        rgtTrkConv[6].Cap[0].dCenterPosConv_cmm := 258800, rgtTrkConv[6].Cap[0].dHeadPos_cmm := 2015800, rgtTrkConv[6].Cap[0].dHeadPosConv_cmm := 388800, rgtTrkConv[6].Cap[0].dPresenceHead_cmm := 2015800, rgtTrkConv[6].Cap[0].dPresenceTail_cmm := 1755800, rgtTrkConv[7].xGlassPresence := 1, rgtTrkConv[7].xPlatePassageNext := 1, rgtTrkConv[7].xGlassPresCom := 1, rgtTrkConv[7].xHeadPresenceConv := 1, rgtTrkConv[7].dStartPosition_cmm := 2127000, rgtTrkConv[7].dEndPosition_cmm := 2627000, rgtTrkConv[7].dStepAdv_cmm[0] := 1620, rgtTrkConv[7].dActualRamp_cmm[0] := 33700, rgtTrkConv[7].dLengthConveyor := 500000, rgtTrkConv[7].dHeadPosition_cmm := 2613400, rgtTrkConv[7].dTailPosition_cmm := 2445700, rgtTrkConv[7].dIndexCaps := 1, rgtTrkConv[7].Cap[0].xHead := 1, rgtTrkConv[7].Cap[0].xCenter := 1, rgtTrkConv[7].Cap[0].xTail := 1, rgtTrkConv[7].Cap[0].xPresence := 1, rgtTrkConv[7].Cap[0].dPointer := 12, rgtTrkConv[7].Cap[0].dTailPos_cmm := 2445700, rgtTrkConv[7].Cap[0].dTailPosConv_cmm := 318700, rgtTrkConv[7].Cap[0].dCenterPos_cmm := 2529550, rgtTrkConv[7].Cap[0].dCenterPosConv_cmm := 402550, rgtTrkConv[7].Cap[0].dHeadPos_cmm := 2613400, rgtTrkConv[7].Cap[0].dHeadPosConv_cmm := 486400, rgtTrkConv[7].Cap[0].dPresenceHead_cmm := 2613400, rgtTrkConv[7].Cap[0].dPresenceTail_cmm := 2445700, rgtTrkConv[8].xPlatePassagePrevious := 1, rgtTrkConv[8].xGlassPresCom := 1, rgtTrkConv[8].dStartPosition_cmm := 2627000, rgtTrkConv[8].dEndPosition_cmm := 2702000, rgtTrkConv[8].dStepAdv_cmm[0] := 1620, rgtTrkConv[8].dActualRamp_cmm[0] := 33700, rgtTrkConv[8].dLengthConveyor := 75000, rgtTrkConv[9].dStartPosition_cmm := 2702000, rgtTrkConv[9].dEndPosition_cmm := 3027000, rgtTrkConv[9].dStepAdv_cmm[0] := 2355, rgtTrkConv[9].dActualRamp_cmm[0] := 33700, rgtTrkConv[9].dLengthConveyor := 325000, rgtTrkConv[10].xGlassPresence := 1, rgtTrkConv[10].xGlassPresCom := 1, rgtTrkConv[10].xHeadPresenceConv := 1, rgtTrkConv[10].dStartPosition_cmm := 3027000, rgtTrkConv[10].dEndPosition_cmm := 3427000, rgtTrkConv[10].dStepAdv_cmm[0] := 2700, rgtTrkConv[10].dActualRamp_cmm[0] := 93700, rgtTrkConv[10].dLengthConveyor := 400000, rgtTrkConv[10].dHeadPosition_cmm := 3312224, rgtTrkConv[10].dTailPosition_cmm := 3052224, rgtTrkConv[10].dIndexCaps := 1, rgtTrkConv[10].Cap[0].xHead := 1, rgtTrkConv[10].Cap[0].xCenter := 1, rgtTrkConv[10].Cap[0].xTail := 1, rgtTrkConv[10].Cap[0].xPresence := 1, rgtTrkConv[10].Cap[0].dPointer := 1, rgtTrkConv[10].Cap[0].dTailPos_cmm := 3052224, rgtTrkConv[10].Cap[0].dTailPosConv_cmm := 25224,
        rgtTrkConv[10].Cap[0].dCenterPos_cmm := 3182224, rgtTrkConv[10].Cap[0].dCenterPosConv_cmm := 155224, rgtTrkConv[10].Cap[0].dHeadPos_cmm := 3312224, rgtTrkConv[10].Cap[0].dHeadPosConv_cmm := 285224, rgtTrkConv[10].Cap[0].dPresenceHead_cmm := 3312224, rgtTrkConv[10].Cap[0].dPresenceTail_cmm := 3052224, rgtTrkConv[11].dStartPosition_cmm := 3427000, rgtTrkConv[11].dEndPosition_cmm := 3777000, rgtTrkConv[11].dStepAdv_cmm[0] := 3000, rgtTrkConv[11].dStepAdv_cmm[1] := 3000, rgtTrkConv[11].dActualRamp_cmm[0] := 93700, rgtTrkConv[11].dActualRamp_cmm[1] := 93700, rgtTrkConv[11].dLengthConveyor := 350000, rgtTrkConv[12].xGlassPresence := 1, rgtTrkConv[12].xPlatePassageNext := 1, rgtTrkConv[12].xGlassPresCom := 1, rgtTrkConv[12].dStartPosition_cmm := 3777000, rgtTrkConv[12].dEndPosition_cmm := 4227000, rgtTrkConv[12].dStepAdv_cmm[0] := 3000, rgtTrkConv[12].dActualRamp_cmm[0] := 93700, rgtTrkConv[12].dLengthConveyor := 450000, rgtTrkConv[12].dTailPosition_cmm := 4202979, rgtTrkConv[12].dIndexCaps := 1, rgtTrkConv[12].Cap[0].xTail := 1, rgtTrkConv[12].Cap[0].xPresence := 1, rgtTrkConv[12].Cap[0].dPointer := 3, rgtTrkConv[12].Cap[0].dTailPos_cmm := 4202979, rgtTrkConv[12].Cap[0].dTailPosConv_cmm := 425979, rgtTrkConv[12].Cap[0].dPresenceHead_cmm := 4370679, rgtTrkConv[12].Cap[0].dPresenceTail_cmm := 4202979, rgtTrkConv[13].xGlassPresence := 1, rgtTrkConv[13].xPlatePassagePrevious := 1, rgtTrkConv[13].xGlassPresCom := 1, rgtTrkConv[13].xHeadPresenceConv := 1, rgtTrkConv[13].dStartPosition_cmm := 4227000, rgtTrkConv[13].dEndPosition_cmm := 4527000, rgtTrkConv[13].dStepAdv_cmm[0] := 3000, rgtTrkConv[13].dStepAdv_cmm[1] := 3000, rgtTrkConv[13].dActualRamp_cmm[0] := 93700, rgtTrkConv[13].dActualRamp_cmm[1] := 93700, rgtTrkConv[13].dLengthConveyor := 300000, rgtTrkConv[13].dHeadPosition_cmm := 4370679, rgtTrkConv[13].dIndexCaps := 1, rgtTrkConv[13].Cap[0].xHead := 1, rgtTrkConv[13].Cap[0].xCenter := 1, rgtTrkConv[13].Cap[0].xPresence := 1, rgtTrkConv[13].Cap[0].dPointer := 3, rgtTrkConv[13].Cap[0].dCenterPos_cmm := 4286829, rgtTrkConv[13].Cap[0].dCenterPosConv_cmm := 59829, rgtTrkConv[13].Cap[0].dHeadPos_cmm := 4370679, rgtTrkConv[13].Cap[0].dHeadPosConv_cmm := 143679, rgtTrkConv[13].Cap[0].dPresenceHead_cmm := 4370679, rgtTrkConv[13].Cap[0].dPresenceTail_cmm := 4202979, rgtTrkConv[14].dStartPosition_cmm := 4527000, rgtTrkConv[14].dEndPosition_cmm := 4627000, rgtTrkConv[14].dStepAdv_cmm[0] := 3300, rgtTrkConv[14].dStepAdv_cmm[1] := 3300, rgtTrkConv[14].dActualRamp_cmm[0] := 93700, rgtTrkConv[14].dActualRamp_cmm[1] := 93700, rgtTrkConv[14].dLengthConveyor := 100000,
        rgtTrkConv[15].dStartPosition_cmm := 4627000, rgtTrkConv[15].dEndPosition_cmm := 5027000, rgtTrkConv[15].dStepAdv_cmm[0] := 2514, rgtTrkConv[15].dActualRamp_cmm[0] := 93700, rgtTrkConv[15].dLengthConveyor := 400000, rgtTrkConv[15].tmON_StopNextConveyor.PRE := 20, rgtTrkConv[16].dStartPosition_cmm := 5027000, rgtTrkConv[16].dEndPosition_cmm := 5427000, rgtTrkConv[16].dStepAdv_cmm[0] := 3300, rgtTrkConv[16].dActualRamp_cmm[0] := 93700, rgtTrkConv[16].dLengthConveyor := 400000, rgtTrkConv[17].dStartPosition_cmm := 5427000, rgtTrkConv[17].dEndPosition_cmm := 5827000, rgtTrkConv[17].dStepAdv_cmm[0] := 2700, rgtTrkConv[17].dActualRamp_cmm[0] := 93700, rgtTrkConv[17].dLengthConveyor := 400000, rgtTrkConv[18].xGlassPresence := 1, rgtTrkConv[18].xPlatePassageNext := 1, rgtTrkConv[18].xGlassPresCom := 1, rgtTrkConv[18].dStartPosition_cmm := 5827000, rgtTrkConv[18].dEndPosition_cmm := 6227000, rgtTrkConv[18].dStepAdv_cmm[0] := 2700, rgtTrkConv[18].dStepAdv_cmm[1] := 2700, rgtTrkConv[18].dActualRamp_cmm[0] := 93700, rgtTrkConv[18].dActualRamp_cmm[1] := 93700, rgtTrkConv[18].dLengthConveyor := 400000, rgtTrkConv[18].dTailPosition_cmm := 6128300, rgtTrkConv[18].dIndexCaps := 1, rgtTrkConv[18].Cap[0].xCenter := 1, rgtTrkConv[18].Cap[0].xTail := 1, rgtTrkConv[18].Cap[0].xPresence := 1, rgtTrkConv[18].Cap[0].dPointer := 8, rgtTrkConv[18].Cap[0].dTailPos_cmm := 6128300, rgtTrkConv[18].Cap[0].dTailPosConv_cmm := 301300, rgtTrkConv[18].Cap[0].dCenterPos_cmm := 6212150, rgtTrkConv[18].Cap[0].dCenterPosConv_cmm := 385150, rgtTrkConv[18].Cap[0].dPresenceHead_cmm := 6296000, rgtTrkConv[18].Cap[0].dPresenceTail_cmm := 6128300, rgtTrkConv[19].xGlassPresence := 1, rgtTrkConv[19].xPlatePassagePrevious := 1, rgtTrkConv[19].xGlassPresCom := 1, rgtTrkConv[19].xHeadPresenceConv := 1, rgtTrkConv[19].dStartPosition_cmm := 6227000, rgtTrkConv[19].dEndPosition_cmm := 6627000, rgtTrkConv[19].dStepAdv_cmm[0] := 2700, rgtTrkConv[19].dActualRamp_cmm[0] := 93700, rgtTrkConv[19].dLengthConveyor := 400000, rgtTrkConv[19].dHeadPosition_cmm := 6296000, rgtTrkConv[19].dIndexCaps := 1, rgtTrkConv[19].Cap[0].xHead := 1, rgtTrkConv[19].Cap[0].xPresence := 1, rgtTrkConv[19].Cap[0].dPointer := 8, rgtTrkConv[19].Cap[0].dHeadPos_cmm := 6296000, rgtTrkConv[19].Cap[0].dHeadPosConv_cmm := 69000, rgtTrkConv[19].Cap[0].dPresenceHead_cmm := 6296000, rgtTrkConv[19].Cap[0].dPresenceTail_cmm := 6128300, rgtTrkConv[20].dStartPosition_cmm := 6627000, rgtTrkConv[20].dEndPosition_cmm := 7027000, rgtTrkConv[20].dStepAdv_cmm[0] := 2700, rgtTrkConv[20].dActualRamp_cmm[0] := 93700,
        rgtTrkConv[20].dLengthConveyor := 400000, rgtTrkConv[21].dStartPosition_cmm := 7027000, rgtTrkConv[21].dEndPosition_cmm := 7427000, rgtTrkConv[21].dStepAdv_cmm[0] := 87, rgtTrkConv[21].dActualRamp_cmm[0] := 93700, rgtTrkConv[21].dLengthConveyor := 400000, rgtTrkConv[22].dStartPosition_cmm := 7427000, rgtTrkConv[22].dEndPosition_cmm := 8177000, rgtTrkConv[22].dStepAdv_cmm[0] := 3000, rgtTrkConv[22].dActualRamp_cmm[0] := 93700, rgtTrkConv[22].dLengthConveyor := 750000, rgtTrkConv[23].dStartPosition_cmm := 8177000, rgtTrkConv[23].dEndPosition_cmm := 8627000, rgtTrkConv[23].dStepAdv_cmm[0] := 3000, rgtTrkConv[23].dActualRamp_cmm[0] := 93700, rgtTrkConv[23].dLengthConveyor := 450000, rgtTrkConv[24].dStartPosition_cmm := 8627000, rgtTrkConv[24].dEndPosition_cmm := 9077000, rgtTrkConv[24].dStepAdv_cmm[0] := 3300, rgtTrkConv[24].dActualRamp_cmm[0] := 93700, rgtTrkConv[24].dLengthConveyor := 450000, rgtTrkConv[25].dStartPosition_cmm := 9077000, rgtTrkConv[25].dEndPosition_cmm := 9372000, rgtTrkConv[25].dStepAdv_cmm[0] := 3300, rgtTrkConv[25].dActualRamp_cmm[0] := 93700, rgtTrkConv[25].dLengthConveyor := 295000, rgtTrkConv[25].tmON_StopNextConveyor.PRE := 20, rgtTrkConv[26].dStartPosition_cmm := 9372000, rgtTrkConv[26].dEndPosition_cmm := 9897000, rgtTrkConv[26].dStepAdv_cmm[0] := 3300, rgtTrkConv[26].dActualRamp_cmm[0] := 93700, rgtTrkConv[26].dLengthConveyor := 525000, rgtTrkConv[26].tmON_StopNextConveyor.PRE := 20, rgtTrkConv[27].dStartPosition_cmm := 9897000, rgtTrkConv[27].dEndPosition_cmm := 10047000, rgtTrkConv[27].dStepAdv_cmm[0] := 2700, rgtTrkConv[27].dActualRamp_cmm[0] := 93700, rgtTrkConv[27].dLengthConveyor := 150000); {access None}
        .rgtTrkConv[6]   // M302M7
        .rgtTrkConv[3]   // M302M4
        .rgtTrkConv[4]   // M302M5
        .rgtTrkConv[7]   // M303M1
        .rgtTrkConv[8]   // M303M2
        .rgtTrkConv[9]   // M304M1
        .rgtTrkConv[10]   // M305M1
        .rgtTrkConv[11]   // M306M1
        .rgtTrkConv[5]   // M302M6
        .rgtTrkConv[0]   // M302M1
        .rgtTrkConv[2]   // M302M3
        .rgtTrkConv[18]   // M307DM1
        .rgtTrkConv[19]   // M307EM1
        .rgtTrkConv[20]   // M307FM1
        .rgtTrkConv[21]   // M350M1
        .rgtTrkConv[1]   // M302M2
        .rgtTrkConv[12]   // M307AM1
        .rgtTrkConv[15]   // M307AM4
        .rgtTrkConv[16]   // M307BM1
        .rgtTrkConv[13]   // M307AM2
        .rgtTrkConv[14]   // M307AM3
        .rgtTrkConv[22]   // M310M1
        .rgtTrkConv[17]   // M307CM1
        .rgtTrkConv[23]   // M310M2
        .rgtTrkConv[24]   // M310M3
        .rgtTrkConv[25]   // M360M1
        .rgtTrkConv[26]   // M315M1
        .rgtTrkConv[27]   // M315M2
        .rgtTrkConv[28]   // M315M3
   Z300_Scada_Continuous : UDT_HMI_LINE_PLATE;
   Z301 : MAC_Zone_ML := (ST_xSelAutoMode := 1, ST_xManualModeConditionOK := 1, ST_xAutoModeAccepted := 1, ST_xConditionOKStopCycle := 1, ST_xCycleON := 1, ST_xConditionOkPhaseAdvancement := 1, ST_xConditionOkCycleON := 1, ST_xEnableControlError := 1, ST_xPLC1 := 1, ST_xThisPlcActive := 1, ST_xConditionOkChangeSpeed := 1, OSR_xThisPlcActive := 1, OSR_xAutoAccepted := 1, INPUT_x24VdcVoltageON := 1, INPUT_xMainEmergencyON := 1, INPUT_xPowerSupply230V_Service := 1, INPUT_xPowerSupply230V_PLC1 := 1, INPUT_xPowerSupply230V_PLC2 := 1, INPUT_xPowerSupply24VLogic1 := 1, INPUT_xPowerSupply24VLogic2 := 1, INPUT_xPowerSupply24VLogic3 := 1, INPUT_xPowerSupply24VDrive1 := 1, INPUT_xPowerSupply24VDrive2 := 1, INPUT_xPowerSupply400VDrive1 := 1, INPUT_xPowerSupply400VDrive2 := 1, INPUT_xPLC_ID_1 := 1, INPUT_xPLC1Selected := 1, INPUT_xEthernetSwitch24VON := 1, OUTPUT_xPLC1Selected := 1, AUX_dLehrSpeed_mm_min := 20336, tmON_ResetAlarm.PRE := 2000, tmON_ResetAlarm.ACC := 2018, tmON_24Vdc.PRE := 2000, tmON_24Vdc.ACC := 2019, tmON_24Vdc.EN := 1, tmON_24Vdc.DN := 1, tmON_400Vca.PRE := 2000, tmON_400Vca.ACC := 2019, tmON_400Vca.EN := 1, tmON_400Vca.DN := 1, tmON_EmergencyOK.PRE := 2000, tmON_EmergencyOK.ACC := 2002, tmON_EmergencyOK.EN := 1, tmON_EmergencyOK.DN := 1, tmON_Cycle.PRE := 15000, tmON_Cycle.ACC := 15000, tmON_Cycle.EN := 1, tmON_Cycle.DN := 1, tmON_ForceStop.PRE := 2000, tmON_AllowStopCleaning.PRE := 10000, tmON_CycleAcousticAlarm.PRE := 15000, tmON_ConveyorsNotOK.PRE := 2000, tmON_StopCycleForFaults.PRE := 2000, tmON_StopCycleForSaturation.PRE := 2000); {access None}
   Z301_ALM : MAC_Zone_ML_ALM; {access Read Only}
        .rgxEmergency[0].0   // Z300.Main emergency stop
        .rgxEmergency[0].1   // Z300.Main emergency stop
        .rgxEmergency[0].2   // Z300.Main emergency stop
        .rgxEmergency[0].3   // Z300.Main emergency stop
        .rgxEmergency[0].31   // MCC1300.Main emergency ON
        .rgxEmergency[0].4   // Z300.Main emergency stop
        .rgxEmergency[0].5   // Z300.Main emergency stop
        .rgxEmergency[0].6   // Z300.Main emergency stop
        .rgxEmergency[0].7   // Z300.Main emergency stop
        .rgxStoppingFault[0].0   // MCC1300.24Vdc Voltage ON
        .rgxStoppingFault[0].13   // MCC1300.Alarm power supply 24V eth switch
        .rgxFault[0].0   // MCC1300.Alarm power supplies 230V PLC1
        .rgxFault[0].1   // MCC1300.Alarm power supplies 230V PLC2
        .rgxStoppingFault[0].25   // MCC1300.Drive power module fault
        .rgxFault[0].8   // MCC1300.Ethernet Switch Fault
        .rgxStoppingFault[0].24   // MCC1300.Drive power module fault
        .rgxStoppingFault[0].8   // MCC1300.Alarm power supply 24V Drive
        .rgxStoppingFault[0].3   // MCC1300.Alarm power supply 24V logic
        .rgxStoppingFault[0].9   // MCC1300.Alarm power supply 24V Drive
        .rgxStoppingFault[0].16   // MCC1300.Alarm power supply 400V Drive
        .rgxStoppingFault[0].4   // MCC1300.Alarm power supply 24V logic
        .rgxStoppingFault[0].17   // MCC1300.Alarm power supply 400V Drive
        .rgxStoppingFault[0].5   // MCC1300.Alarm power supply 24V logic
   Z301_HMR : MAC_Zone_ML_HMR := (xAutoSpeedAdjustEnabled := 1, dZoneMode := 4, dZoneState := 1, dCleaningState := 2, dAutoSpeedForBreakings_mm_min := 54000, dAutoSpeed_mm_min := 90000, dManualSpeed_mm_min := 20000, dMinAutoSpeedForBreakings_mm_min := 54000, dMinAutoSpeed_mm_min := 90000, rSpeedRatioBreakings := 3.5, rSpeedRatio := 3.0); {access Read Only}
        .rgxMan.0   // Forward all (zone)
        .rgxMan.1   // Backward all (zone)
        .rgxMan.2   // Forward all (line)
        .rgxMan.3   // Backward all (line)
   Z301_HMW : MAC_Zone_ML_HMW := (xEnDisableAutoSpeedAdjust := 1, dAutoSpeedForBreakings_mm_min := 54000, dAutoSpeed_mm_min := 90000, dManualSpeed_mm_min := 20000, rSpeedRatioBreakings := 3.0, rSpeedRatio := 3.0);
        .rgxMan.0   // Forward all (zone) {x|x|x|x|O}
        .rgxMan.1   // Backward all (zone) {x|x|x|x|O}
        .rgxMan.2   // Forward all (line) {x|x|x|x|O}
        .rgxMan.3   // Backward all (line) {x|x|x|x|O}
   Z311S : MAC_SafetyAccess; {access Read Only}
   Z311S_ALM : MAC_SafetyAccess_ALM;
        .rgxFault[0].0   // Z401.M311S.Safety area intervened
        .rgxFault[0].1   // Z401.M311S.Door open
   Z311S_HMR : MAC_SafetyAccess_HMR; {access Read Only}
   Z311S_INPUT_xAccessReqRotator : BOOL; {access Read Only}
   Z311S_INPUT_xSafetyAreaRotator : BOOL; {access Read Only}
   Z311S_OUTPUT_xEL_AccessAcceptedRotator : BOOL; {access Read Only}
   Z311S_OUTPUT_xHL_AccessAcceptedRotator : BOOL; {access Read Only}
   Z311S_OUTPUT_xHL_SafetyAreaRotatorNOK : BOOL; {access Read Only}
   Z316S : MAC_SafetyAccess; {access Read Only}
   Z316S_ALM : MAC_SafetyAccess_ALM;
        .rgxFault[0].0   // Z402.M316S.Safety area intervened
        .rgxFault[0].1   // Z402.M316S.Door open
   Z316S_HMR : MAC_SafetyAccess_HMR; {access Read Only}
   Z316S_INPUT_xAccessReqRotator : BOOL; {access Read Only}
   Z316S_INPUT_xSafetyAreaRotator : BOOL; {access Read Only}
   Z316S_OUTPUT_xEL_AccessAcceptedRotator : BOOL; {access Read Only}
   Z316S_OUTPUT_xHL_AccessAcceptedRotator : BOOL; {access Read Only}
   Z316S_OUTPUT_xHL_SafetyAreaRotatorNOK : BOOL; {access Read Only}
   Z401 : MAC_Zone := (ST_xCycleON := 1, ST_xConditionOkPhaseAdvancement := 1, ST_xConditionOkCycleON := 1, ST_xCleaningConditionOK := 1, ST_xAutoModeAccepted := 1, ST_xSelectionAutomaticMode := 1, ST_xEnableControlError := 1, OSR_xAutomaticMode := 1, AUX_dSpeedStandby_mm_min := 12000, AUX_dSpeedTINUnload_mm_min := 81000, AUX_dProgressiveID := 356828, tmON_ResetAlarm.PRE := 1000, tmON_ResetAlarm.ACC := 1000, tmON_24Vdc.PRE := 2000, tmON_24Vdc.ACC := 2000, tmON_24Vdc.EN := 1, tmON_24Vdc.DN := 1, tmON_400Vca.PRE := 2000, tmON_400Vca.ACC := 2019, tmON_400Vca.EN := 1, tmON_400Vca.DN := 1, tmON_EmergencyOK.PRE := 2000, tmON_EmergencyOK.ACC := 2000, tmON_EmergencyOK.EN := 1, tmON_EmergencyOK.DN := 1, tmON_Cycle.PRE := 15000, tmON_Cycle.ACC := 15000, tmON_Cycle.EN := 1, tmON_Cycle.DN := 1, tmON_ForceStop.PRE := 2000, tmON_CycleAcousticAlarm.PRE := 10000); {access None}
   Z401_ALM : MAC_Zone_ALM;
        .rgxFault[0].0   // Z400.MCC1401.24Vdc Voltage
        .rgxFault[0].6   // Z400.MCC1401.P18QF2.Alarm power supply 24V logic
        .rgxFault[0].7   // Z400.MCC1401.P18QF3.Alarm power supply 24V logic
        .rgxFault[0].8   // Z400.MCC1401.P19QF1.Alarm power supply 24V logic
        .rgxFault[0].9   // Z400.MCC1401.P155SW1.Ethernet switch power supply
        .rgxStoppingFault[0].0   // Z400.P41GS1.Power module 1 Fault
        .rgxEmergency[0].1   // Z401.MCC1401.General emergency ON
        .rgxEmergency[0].10   // Z401.CS4401.Emergency localization
        .rgxEmergency[0].8   // Z401.M311S.Emergency localization
        .rgxEmergency[0].9   // Z401.M311S.Emergency localization
        .rgxWarning[0].0   // Z400.MCC1401.P20QF3.Alarm power supply 24V drives
        .rgxWarning[0].1   // Z400.MCC1401.P11QF2/P11QF1D/P11QF1.Alarm power supplies 230Vac cabinet
        .rgxWarning[0].3   // Z400.MCC1401.P41QM1.Drive power module supply
        .rgxWarning[0].4   // Z400.MCC1401.P11QF4.Alarm power supplies 230Vac cabinet
   Z401_HMI_rgtPlateScada : HMI_LiteData[5,2,7] := ([3,0,0].dHead_PosX_mm := 3200, [3,0,0].dTail_PosX_mm := 1400, [3,0,0].dPlateLength_mm := 1800, [3,0,0].dPositionY_mm := 250, [3,0,0].dPlateWidth_mm := 2600, [3,0,0].dPlateId := 3658556, [3,0,0].dProductionID := 1029, [3,0,0].dDestination := 3, [3,0,0].dAlternative := 4);
        [0,0,0]   // M310B
        [1,0,0]   // M310A
        [2,0,0]   // M311
        [3,0,0]   // M311A
        [4,0,0]   // M312
   Z401_HMI_rgtPlateScada_Internal : HMI_LiteData[5,2,7] := ([3,0,0].dHead_PosX_mm := 3200, [3,0,0].dTail_PosX_mm := 1400, [3,0,0].dPlateLength_mm := 1800, [3,0,0].dPositionY_mm := 250, [3,0,0].dPlateWidth_mm := 2600, [3,0,0].dPlateId := 3658556, [3,0,0].dProductionID := 1029, [3,0,0].dDestination := 3, [3,0,0].dAlternative := 4);
        [0,0,0]   // M310B
        [1,0,0]   // M310A
        [2,0,0]   // M311
        [3,0,0]   // M311A
        [4,0,0]   // M312
   Z401_HMR : MAC_Zone_HMR := (dZoneMode := 4, dZoneState := 1, dCleaningState := 2, dLineSpeed_mm_min := 60000);
        .rgxMan.0   // Forward alll
        .rgxMan.1   // Backward all
   Z401_HMW : MAC_Zone_HMW := (dLocalRemoteSettings := 1, dLineSpeed_mm_min := 60000, dManualSpeed_mm_min := 60000);
        .rgxMan.0   // Forward alll
        .rgxMan.1   // Backward all
   Z401_INPUT_xMainLineEmergencyON : BOOL; {access Read Only}
   Z401_OUTPUT_xMCC_SafetyPanel1 : BOOL; {access Read Only}
   Z401S_INPUT_xSafetyAreaPopup : BOOL; {access Read Only}
   Z401S_INPUT_xSafetyAreaRotator : BOOL; {access Read Only}
   Z402 : MAC_Zone := (ST_xCycleON := 1, ST_xConditionOkPhaseAdvancement := 1, ST_xConditionOkCycleON := 1, ST_xCleaningConditionOK := 1, ST_xAutoModeAccepted := 1, ST_xSelectionAutomaticMode := 1, ST_xEnableControlError := 1, OSR_xAutomaticMode := 1, AUX_dSpeedStandby_mm_min := 12000, AUX_dSpeedTINUnload_mm_min := 81000, AUX_dProgressiveID := 356828, tmON_ResetAlarm.PRE := 1000, tmON_ResetAlarm.ACC := 1000, tmON_24Vdc.PRE := 2000, tmON_24Vdc.ACC := 2000, tmON_24Vdc.EN := 1, tmON_24Vdc.DN := 1, tmON_400Vca.PRE := 2000, tmON_400Vca.ACC := 2019, tmON_400Vca.EN := 1, tmON_400Vca.DN := 1, tmON_EmergencyOK.PRE := 2000, tmON_EmergencyOK.ACC := 2000, tmON_EmergencyOK.EN := 1, tmON_EmergencyOK.DN := 1, tmON_Cycle.PRE := 15000, tmON_Cycle.ACC := 15000, tmON_Cycle.EN := 1, tmON_Cycle.DN := 1, tmON_ForceStop.PRE := 2000, tmON_CycleAcousticAlarm.PRE := 10000); {access None}
   Z402_ALM : MAC_Zone_ALM;
        .rgxFault[0].0   // Z400.MCC1401.24Vdc Voltage
        .rgxFault[0].6   // Z400.MCC1401.P18QF2.Alarm power supply 24V logic
        .rgxFault[0].7   // Z400.MCC1401.P18QF3.Alarm power supply 24V logic
        .rgxFault[0].8   // Z400.MCC1401.P19QF1.Alarm power supply 24V logic
        .rgxFault[0].9   // Z400.MCC1401.P155SW1.Ethernet switch power supply
        .rgxStoppingFault[0].0   // Z400.P41GS1.Power module 1 Fault
        .rgxEmergency[0].1   // Z402.MCC1402.General emergency ON
        .rgxEmergency[0].10   // Z402.CS4402.Emergency localization
        .rgxEmergency[0].8   // Z402.M316S.Emergency localization
        .rgxEmergency[0].9   // Z402.M316S.Emergency localization
        .rgxWarning[0].0   // Z400.MCC1401.P20QF3.Alarm power supply 24V drives
        .rgxWarning[0].1   // Z400.MCC1401.P11QF2/P11QF1D/P11QF1.Alarm power supplies 230Vac cabinet
        .rgxWarning[0].3   // Z400.MCC1401.P41QM1.Drive power module supply
        .rgxWarning[0].4   // Z400.MCC1401.P11QF4.Alarm power supplies 230Vac cabinet
   Z402_HMI_rgtPlateScada : HMI_LiteData[5,2,7] := ([3,0,0].dHead_PosX_mm := 3200, [3,0,0].dTail_PosX_mm := 1400, [3,0,0].dPlateLength_mm := 1800, [3,0,0].dPositionY_mm := 250, [3,0,0].dPlateWidth_mm := 2600, [3,0,0].dPlateId := 3658556, [3,0,0].dProductionID := 1029, [3,0,0].dDestination := 3, [3,0,0].dAlternative := 4);
        [0,0,0]   // M315B
        [1,0,0]   // M315A
        [2,0,0]   // M316
        [3,0,0]   // M316A
        [4,0,0]   // M317
   Z402_HMI_rgtPlateScada_Internal : HMI_LiteData[5,2,7] := ([3,0,0].dHead_PosX_mm := 3200, [3,0,0].dTail_PosX_mm := 1400, [3,0,0].dPlateLength_mm := 1800, [3,0,0].dPositionY_mm := 250, [3,0,0].dPlateWidth_mm := 2600, [3,0,0].dPlateId := 3658556, [3,0,0].dProductionID := 1029, [3,0,0].dDestination := 3, [3,0,0].dAlternative := 4);
        [0,0,0]   // M315B
        [1,0,0]   // M315A
        [2,0,0]   // M316
        [3,0,0]   // M316A
        [4,0,0]   // M317
   Z402_HMR : MAC_Zone_HMR := (dZoneMode := 4, dZoneState := 1, dCleaningState := 2, dLineSpeed_mm_min := 60000);
        .rgxMan.0   // Forward alll
        .rgxMan.1   // Backward all
   Z402_HMW : MAC_Zone_HMW := (dLocalRemoteSettings := 1, dLineSpeed_mm_min := 60000, dManualSpeed_mm_min := 60000);
        .rgxMan.0   // Forward alll
        .rgxMan.1   // Backward all
   Z402_INPUT_xMainLineEmergencyON : BOOL; {access Read Only}
   Z402_OUTPUT_xMCC_SafetyPanel : BOOL; {access Read Only}
   Z402_OUTPUT_xMCC_SafetyPanel1 : BOOL; {access Read Only}
   Z402S_INPUT_xSafetyAreaPopup : BOOL; {access Read Only}
   Z402S_INPUT_xSafetyAreaRotator : BOOL; {access Read Only}
   Z900 : MAC_Zone := (ST_xConditionOKStopCycle := 1, ST_xCycleON := 1, ST_xConditionOkPhaseAdvancement := 1, ST_xConditionOkCycleON := 1, ST_xConditionOkManualMode := 1, ST_xAutoModeAccepted := 1, ST_xSelectionAutomaticMode := 1, ST_xEnableControlError := 1, OSR_xAutomaticMode := 1, AUX_dSpeedStandby_mm_min := 12000, AUX_dSpeedTINUnload_mm_min := 81000, AUX_dProgressiveID := 356828, tmON_ResetAlarm.PRE := 1000, tmON_ResetAlarm.ACC := 1000, tmON_24Vdc.PRE := 2000, tmON_24Vdc.ACC := 2000, tmON_24Vdc.EN := 1, tmON_24Vdc.DN := 1, tmON_400Vca.PRE := 2000, tmON_400Vca.ACC := 2019, tmON_400Vca.EN := 1, tmON_400Vca.DN := 1, tmON_EmergencyOK.PRE := 2000, tmON_EmergencyOK.ACC := 2000, tmON_EmergencyOK.EN := 1, tmON_EmergencyOK.DN := 1, tmON_Cycle.PRE := 3000, tmON_Cycle.ACC := 3000, tmON_Cycle.EN := 1, tmON_Cycle.DN := 1, tmON_ForceStop.PRE := 2000, tmON_CycleAcousticAlarm.PRE := 10000); {access None}
   Z900_ALM : MAC_Zone_ALM;
   Z900_HMI_rgtPlateScada : HMI_LiteData[5,2,7];
        [3,0,0]   // Spare
        [4,0,0]   // Spare
        [0,0,0]   // M351
        [1,0,0]   // M352
        [2,0,0]   // M353
   Z900_HMI_rgtPlateScada_Internal : HMI_LiteData[5,2,7];
        [3,0,0]   // Spare
        [4,0,0]   // Spare
        [0,0,0]   // M351
        [1,0,0]   // M352
        [2,0,0]   // M353
   Z900_HMR : MAC_Zone_HMR := (dZoneMode := 4, dZoneState := 1, dCleaningState := 2, dLineSpeed_mm_min := 50000, dSnapSpeed_mm_min := 8000);
        .rgxMan.0   // Forward alll
        .rgxMan.1   // Backward all
   Z900_HMW : MAC_Zone_HMW := (dLocalRemoteSettings := 1, dLineSpeed_mm_min := 50000, dSnapSpeed_mm_min := 10583, dManualSpeed_mm_min := 21000);
        .rgxMan.0   // Forward alll
        .rgxMan.1   // Backward all
END_VAR

PROGRAM _18_STI   (* main routine _18_STI *)

ROUTINE _18_STI   (* ladder *)
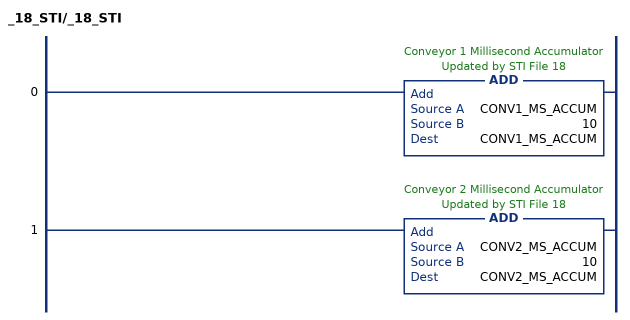
   0: ADD(CONV1_MS_ACCUM,10,CONV1_MS_ACCUM);
   1: ADD(CONV2_MS_ACCUM,10,CONV2_MS_ACCUM);
END_ROUTINE
END_PROGRAM

PROGRAM CommandLogic   (* main routine Main *)

ROUTINE M302M1_Conveyor_Output   (* ladder *)
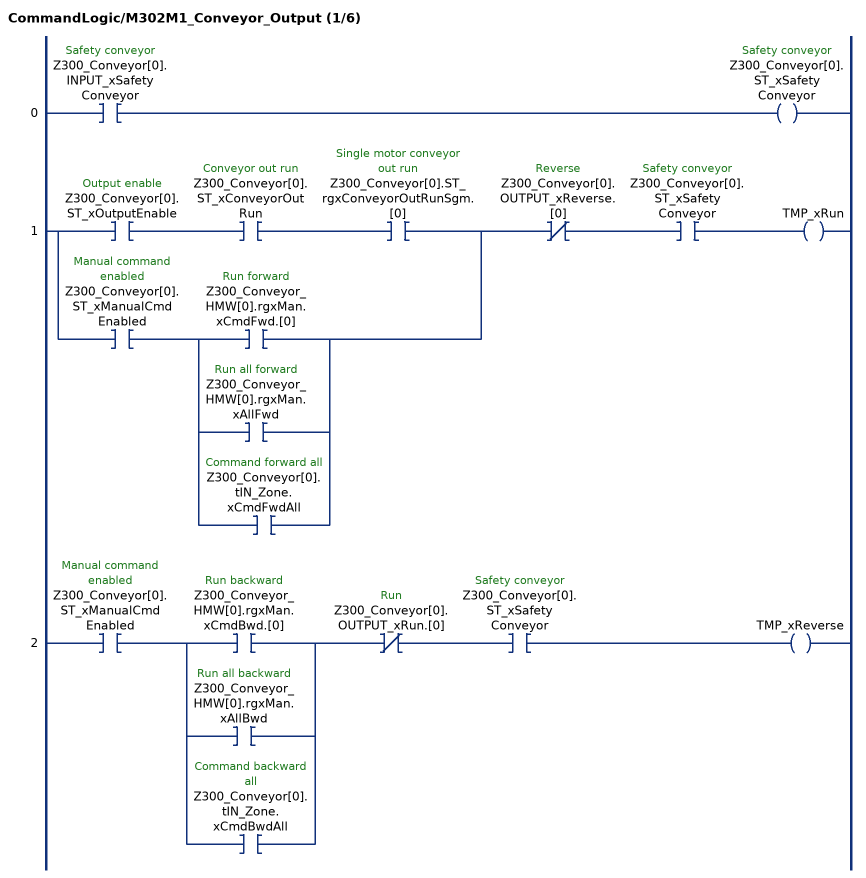
   0: XIC(Z300_Conveyor[0].INPUT_xSafetyConveyor)OTE(Z300_Conveyor[0].ST_xSafetyConveyor);
   1: [XIC(Z300_Conveyor[0].ST_xOutputEnable) XIC(Z300_Conveyor[0].ST_xConveyorOutRun) XIC(Z300_Conveyor[0].ST_rgxConveyorOutRunSgm.[0]) ,XIC(Z300_Conveyor[0].ST_xManualCmdEnabled) [XIC(Z300_Conveyor_HMW[0].rgxMan.xCmdFwd.[0]) ,XIC(Z300_Conveyor_HMW[0].rgxMan.xAllFwd) ,XIC(Z300_Conveyor[0].tIN_Zone.xCmdFwdAll) ] ]XIO(Z300_Conveyor[0].OUTPUT_xReverse.[0])XIC(Z300_Conveyor[0].ST_xSafetyConveyor)OTE(TMP_xRun);
   2: XIC(Z300_Conveyor[0].ST_xManualCmdEnabled)[XIC(Z300_Conveyor_HMW[0].rgxMan.xCmdBwd.[0]) ,XIC(Z300_Conveyor_HMW[0].rgxMan.xAllBwd) ,XIC(Z300_Conveyor[0].tIN_Zone.xCmdBwdAll) ]XIO(Z300_Conveyor[0].OUTPUT_xRun.[0])XIC(Z300_Conveyor[0].ST_xSafetyConveyor)OTE(TMP_xReverse);
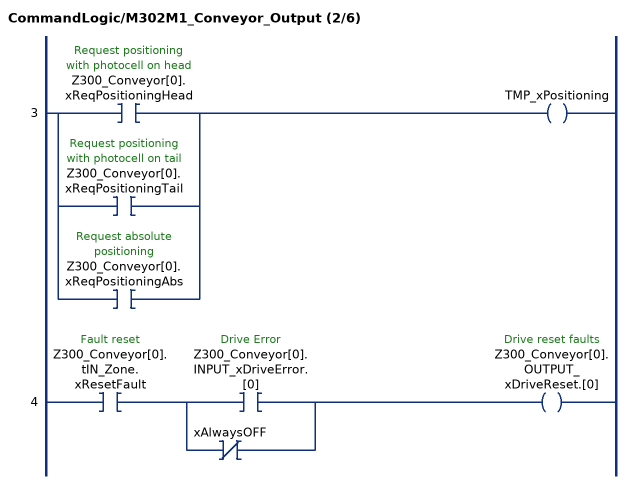
   3: [XIC(Z300_Conveyor[0].xReqPositioningHead) ,XIC(Z300_Conveyor[0].xReqPositioningTail) ,XIC(Z300_Conveyor[0].xReqPositioningAbs) ]OTE(TMP_xPositioning);
   4: XIC(Z300_Conveyor[0].tIN_Zone.xResetFault)[XIC(Z300_Conveyor[0].INPUT_xDriveError.[0]) ,XIO(xAlwaysOFF) ]OTE(Z300_Conveyor[0].OUTPUT_xDriveReset.[0]);
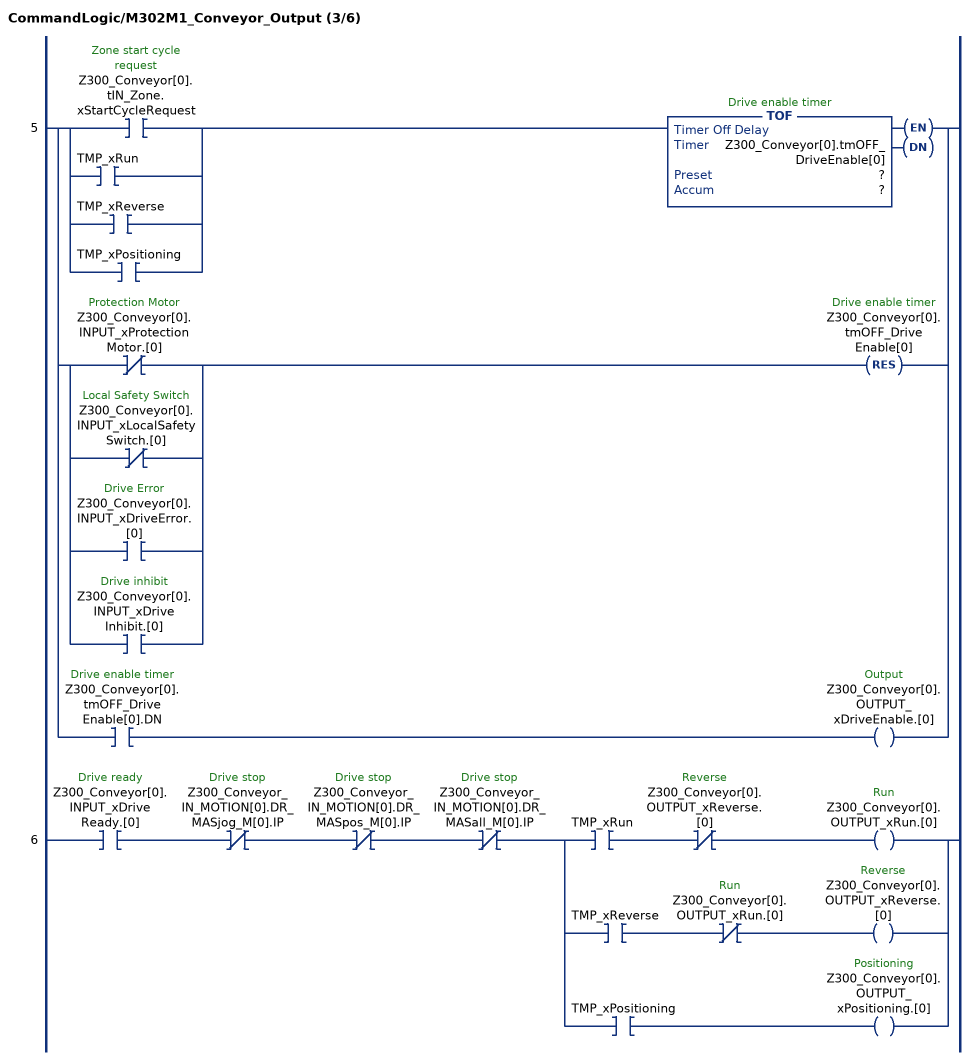
   5: [[XIC(Z300_Conveyor[0].tIN_Zone.xStartCycleRequest) ,XIC(TMP_xRun) ,XIC(TMP_xReverse) ,XIC(TMP_xPositioning) ] TOF(Z300_Conveyor[0].tmOFF_DriveEnable[0],?,?) ,[XIO(Z300_Conveyor[0].INPUT_xProtectionMotor.[0]) ,XIO(Z300_Conveyor[0].INPUT_xLocalSafetySwitch.[0]) ,XIC(Z300_Conveyor[0].INPUT_xDriveError.[0]) ,XIC(Z300_Conveyor[0].INPUT_xDriveInhibit.[0]) ] RES(Z300_Conveyor[0].tmOFF_DriveEnable[0]) ,XIC(Z300_Conveyor[0].tmOFF_DriveEnable[0].DN) OTE(Z300_Conveyor[0].OUTPUT_xDriveEnable.[0]) ];
   6: XIC(Z300_Conveyor[0].INPUT_xDriveReady.[0])XIO(Z300_Conveyor_IN_MOTION[0].DR_MASjog_M[0].IP)XIO(Z300_Conveyor_IN_MOTION[0].DR_MASpos_M[0].IP)XIO(Z300_Conveyor_IN_MOTION[0].DR_MASall_M[0].IP)[XIC(TMP_xRun) XIO(Z300_Conveyor[0].OUTPUT_xReverse.[0]) OTE(Z300_Conveyor[0].OUTPUT_xRun.[0]) ,XIC(TMP_xReverse) XIO(Z300_Conveyor[0].OUTPUT_xRun.[0]) OTE(Z300_Conveyor[0].OUTPUT_xReverse.[0]) ,XIC(TMP_xPositioning) OTE(Z300_Conveyor[0].OUTPUT_xPositioning.[0]) ];
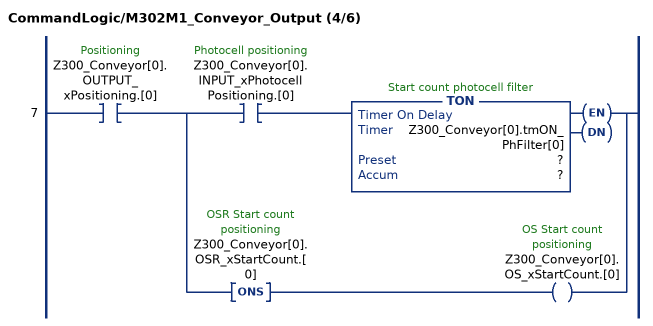
   7: XIC(Z300_Conveyor[0].OUTPUT_xPositioning.[0])[XIC(Z300_Conveyor[0].INPUT_xPhotocellPositioning.[0]) TON(Z300_Conveyor[0].tmON_PhFilter[0],?,?) ,ONS(Z300_Conveyor[0].OSR_xStartCount.[0]) OTE(Z300_Conveyor[0].OS_xStartCount.[0]) ];
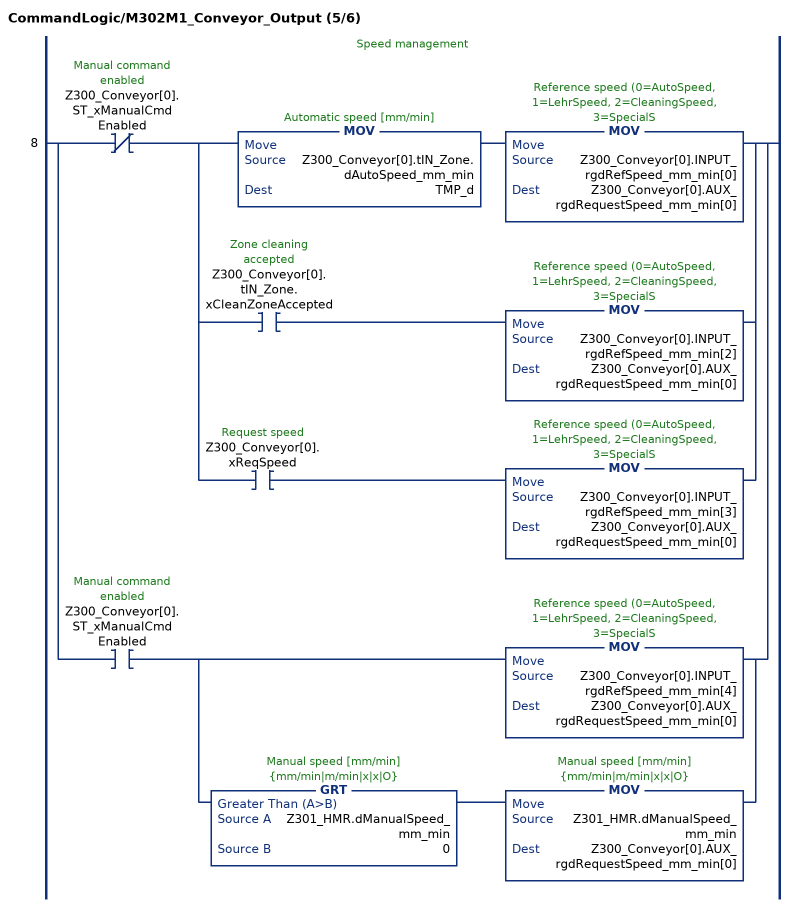
   // Speed management
   8: [XIO(Z300_Conveyor[0].ST_xManualCmdEnabled) [MOV(Z300_Conveyor[0].tIN_Zone.dAutoSpeed_mm_min,TMP_d) MOV(Z300_Conveyor[0].INPUT_rgdRefSpeed_mm_min[0],Z300_Conveyor[0].AUX_rgdRequestSpeed_mm_min[0]) ,XIC(Z300_Conveyor[0].tIN_Zone.xCleanZoneAccepted) MOV(Z300_Conveyor[0].INPUT_rgdRefSpeed_mm_min[2],Z300_Conveyor[0].AUX_rgdRequestSpeed_mm_min[0]) ,XIC(Z300_Conveyor[0].xReqSpeed) MOV(Z300_Conveyor[0].INPUT_rgdRefSpeed_mm_min[3],Z300_Conveyor[0].AUX_rgdRequestSpeed_mm_min[0]) ] ,XIC(Z300_Conveyor[0].ST_xManualCmdEnabled) [MOV(Z300_Conveyor[0].INPUT_rgdRefSpeed_mm_min[4],Z300_Conveyor[0].AUX_rgdRequestSpeed_mm_min[0]) ,GRT(Z301_HMR.dManualSpeed_mm_min,0) MOV(Z301_HMR.dManualSpeed_mm_min,Z300_Conveyor[0].AUX_rgdRequestSpeed_mm_min[0]) ] ];
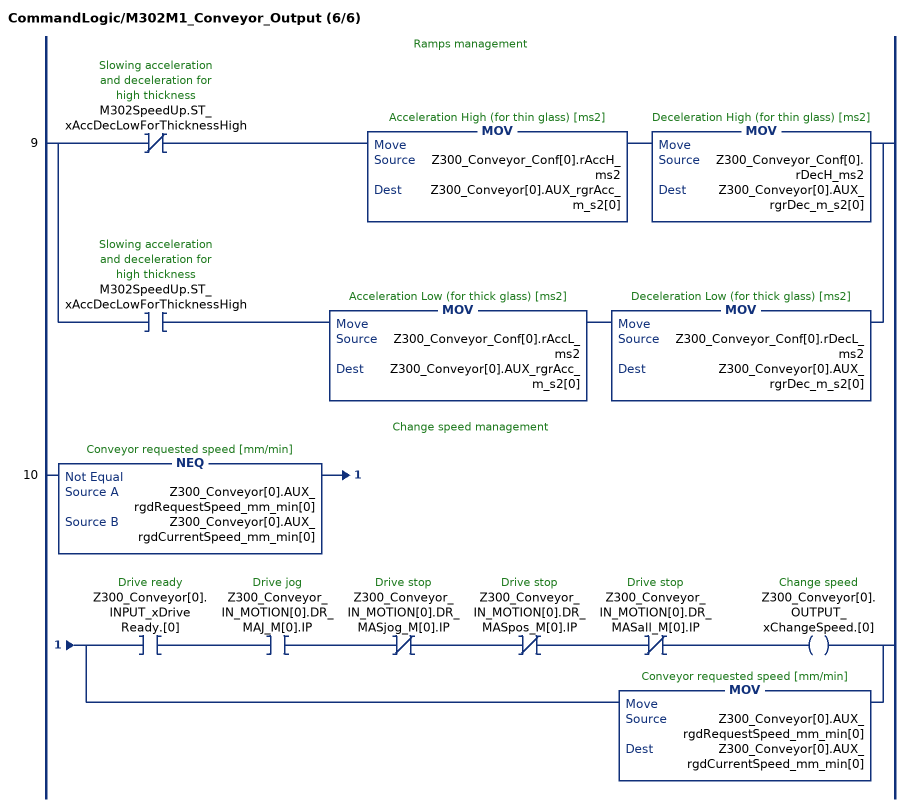
   // Ramps management
   9: [XIO(M302SpeedUp.ST_xAccDecLowForThicknessHigh) MOV(Z300_Conveyor_Conf[0].rAccH_ms2,Z300_Conveyor[0].AUX_rgrAcc_m_s2[0]) MOV(Z300_Conveyor_Conf[0].rDecH_ms2,Z300_Conveyor[0].AUX_rgrDec_m_s2[0]) ,XIC(M302SpeedUp.ST_xAccDecLowForThicknessHigh) MOV(Z300_Conveyor_Conf[0].rAccL_ms2,Z300_Conveyor[0].AUX_rgrAcc_m_s2[0]) MOV(Z300_Conveyor_Conf[0].rDecL_ms2,Z300_Conveyor[0].AUX_rgrDec_m_s2[0]) ];
   // Change speed management
   10: NEQ(Z300_Conveyor[0].AUX_rgdRequestSpeed_mm_min[0],Z300_Conveyor[0].AUX_rgdCurrentSpeed_mm_min[0])[XIC(Z300_Conveyor[0].INPUT_xDriveReady.[0]) XIC(Z300_Conveyor_IN_MOTION[0].DR_MAJ_M[0].IP) XIO(Z300_Conveyor_IN_MOTION[0].DR_MASjog_M[0].IP) XIO(Z300_Conveyor_IN_MOTION[0].DR_MASpos_M[0].IP) XIO(Z300_Conveyor_IN_MOTION[0].DR_MASall_M[0].IP) OTE(Z300_Conveyor[0].OUTPUT_xChangeSpeed.[0]) ,MOV(Z300_Conveyor[0].AUX_rgdRequestSpeed_mm_min[0],Z300_Conveyor[0].AUX_rgdCurrentSpeed_mm_min[0]) ];
END_ROUTINE
